
           // check axes state
           FOR #tempAxisCtr := 1 TO #MAX_NO_OF_AXES DO
             // check for axes to be existing
             IF #statAxes[#tempAxisCtr].typeOfAxis <> #AXIS_NOT_USED THEN
               // check type of axes used
               IF #statAxes[#tempAxisCtr].typeOfAxis = #TYPE_POSITIONING_AXIS THEN
                 // read TO_PositioningAxis status word
                 "LKinCtrl_GetPosAxisData"(posAxis := #statAxes[#tempAxisCtr].axis,
                                           statusWord => #statAxisStatusWord,
                                           errorDetailNumber => #statAxisErrorDetailNumber);
               ELSIF #statAxes[#tempAxisCtr].typeOfAxis = #TYPE_SYNCHRONOUS_AXIS THEN
                 // read TO_SynchronousAxis status word
                 "LKinCtrl_GetSyncAxisData"(syncAxis := #statAxes[#tempAxisCtr].axis,
                                            statusWord => #statAxisStatusWord,
                                            errorDetailNumber => #statAxisErrorDetailNumber);
               END_IF;
             END_IF;

             IF #statAxisStatusWord.%X1 = FALSE THEN
               // do nothing here, continue checks
               ;
             ELSE
               // set status
               #statStatus := #ERR_AXIS_ERROR;
               // set error bit
               #statErrorAutoCleared := TRUE;
               // write axis number to diagnostics
               #statAxisNumberDiag := #tempAxisCtr;
               // set subFunctionStatus
               #statErrorDetailNumber := #statAxisErrorDetailNumber;
               // go to error state
               #statStateMachine := #ERROR_STATE;
               EXIT;
             END_IF;

           END_FOR;

         END_REGION ENABLED_AXES


       #DISABLING_AXES: // Disabling active
         REGION DISABLING_AXES
           // set status message
           #statStatus := #STATUS_DISABLING_AXES_IN_PROGRESS;

           FOR #tempAxisCtr := 1 TO #MAX_NO_OF_AXES DO
             // check for axes to be existing
             IF #statAxes[#tempAxisCtr].typeOfAxis <> #AXIS_NOT_USED THEN
               // set execute trigger for MC_POWER
               #statEnableAxis[#tempAxisCtr] := FALSE;
             END_IF;
           END_FOR;

           // reset enabled axes counter
           #statDisabledAxesCtr := 0;
           // check for disabling to have completed successfully
           FOR #tempAxisCtr := 1 TO #MAX_NO_OF_AXES DO
             // only run code for existing axes
             IF #statAxes[#tempAxisCtr].typeOfAxis <> #AXIS_NOT_USED THEN
               // check for disabling to be done
               IF #instMC_Power[#tempAxisCtr].Status = FALSE THEN
                 // count done signals
                 #statDisabledAxesCtr += 1;
               ELSIF #instMC_Power[#tempAxisCtr].Error THEN
                 // set status
                 #statStatus := #ERR_MC_POWER;
                 // set error bit
                 #statErrorAutoCleared := TRUE;
                 // write MC_HOME errorID to diagnostics
                 #statSubfunctionStatus := #instMC_Power[#tempAxisCtr].ErrorId;
                 // write axis number to diagnostics
                 #statAxisNumberDiag := #tempAxisCtr;
                 // exit FOR loop once error is found
                 EXIT;
                 // go to error state
                 #statStateMachine := #ERROR_STATE;
               END_IF;
             END_IF;
           END_FOR;

           // check for all axes to be enabled successfully
           IF #statDisabledAxesCtr = #statExsitingAxesCtr THEN
             // set status message
             #statStatus := #STATUS_ALL_AXES_DISABLED;
             // reset variable for axesEnabled output
             #statAxesEnabled := FALSE;
             // go to next state
             #statStateMachine := #DISABLED_AXES;
           END_IF;
         END_REGION DISABLING_AXES

       #DISABLED_AXES:
         REGION DISABLED_AXES
           // when disabling is complete the bit #statDisablingCompleted must be set
           #statDisablingCompleted := TRUE;
         END_REGION DISABLED_AXES


       #ERROR_STATE:
         REGION ERROR_STATE
           // Reset axesEnabled output in case of error
           #statAxesEnabled := FALSE;
         END_REGION ERROR_STATE

       ELSE // Undefined state in state machine reached
         #statStatus := #ERR_UNDEFINED_STATE;
         #statErrorUserCleared := TRUE;
     END_CASE;
   END_REGION STATE_MACHINE


   REGION CALL_MC_POWER

     FOR #tempAxisCtr := 1 TO #MAX_NO_OF_AXES DO
       // check for axes to be existing
       IF #statAxes[#tempAxisCtr].typeOfAxis <> #AXIS_NOT_USED THEN
         // check for used axis type to call corresponding FCs
         IF #statAxes[#tempAxisCtr].typeOfAxis = #TYPE_POSITIONING_AXIS THEN
           // call MC_HOME for available positioning axes
           "LKinCtrl_CallMC_Power_PosAxis"(posAxisIn := #statAxes[#tempAxisCtr].axis,
                                           enable := #statEnableAxis[#tempAxisCtr],
                                           startMode := #startMode[#tempAxisCtr],
                                           stopMode := #stopMode[#tempAxisCtr],
                                           instMC_Power := #instMC_Power[#tempAxisCtr]);
           // check for error to be pending
           IF #instMC_Power[#tempAxisCtr].Error
             // check for no axis or kinematics errors detected prior
             AND #statStatus <> #ERR_AXIS_ERROR
             AND #statStatus <> #ERR_KIN_ERROR
           THEN
             // set status
             #statStatus := #ERR_MC_POWER;
             // set error bit
             #statErrorAutoCleared := TRUE;
             // write MC_HOME errorID to diagnostics
             #statSubfunctionStatus := #instMC_Power[#tempAxisCtr].ErrorId;
             // write axis number to diagnostics
             #statAxisNumberDiag := #tempAxisCtr;
             // exit FOR loop once error is found
             EXIT;
             // go to error state
             #statStateMachine := #ERROR_STATE;
           END_IF;

         ELSIF #statAxes[#tempAxisCtr].typeOfAxis = #TYPE_SYNCHRONOUS_AXIS THEN
           // call MC_HOME for available synchronous axes
           "LKinCtrl_CallMC_Power_SyncAxis"(syncAxisIn := #statAxes[#tempAxisCtr].axis,
                                            enable := #statEnableAxis[#tempAxisCtr],
                                            startMode := #startMode[#tempAxisCtr],
                                            stopMode := #stopMode[#tempAxisCtr],
                                            instMC_Power := #instMC_Power[#tempAxisCtr]);
           // check for error to be pending
           IF #instMC_Power[#tempAxisCtr].Error
             // check for no axis or kinematics errors detected prior
             AND #statStatus <> #ERR_AXIS_ERROR
             AND #statStatus <> #ERR_KIN_ERROR
           THEN
             // set status
             #statStatus := #ERR_MC_POWER;
             // set error bit
             #statErrorAutoCleared := TRUE;
             // write MC_HOME errorID to diagnostics
             #statSubfunctionStatus := #instMC_Power[#tempAxisCtr].ErrorId;
             // write axis number to diagnostics
             #statAxisNumberDiag := #tempAxisCtr;
             // exit FOR loop once error is found
             EXIT;
             // go to error state
             #statStateMachine := #ERROR_STATE;
           END_IF;
         END_IF;

       END_IF;
     END_FOR;

   END_REGION CALL_MC_POWER


   REGION OUTPUTS
     // Write outputs
     IF (#statDisablingCompleted = TRUE) THEN
       // Reset outputs if disabling completed
       #statBusy := FALSE;
       #statError := FALSE;
       #statErrorUserCleared := FALSE;
       #statErrorAutoCleared := FALSE;
       #statStatus := #STATUS_NO_CALL;
       #statStateMachine := #NO_PROCESSING; // Switch state machine to "no processing"

     ELSIF (#statErrorUserCleared = TRUE) AND (#statError = FALSE) THEN
       // Error can only be cleared by user; rising edge at enable input is needed to continue 
       #statBusy := FALSE;
       #statError := TRUE;
       #statStateMachine := #NO_PROCESSING; // Switch state machine to "no processing"

     ELSIF (#statErrorAutoCleared = TRUE) AND (#statError = FALSE) THEN
       // Error can be reset by FB automatically  
       #statBusy := TRUE;
       #statError := TRUE;
       // TODO: Handling of autocleared error

     ELSIF (#statErrorAutoCleared = FALSE) AND (#statErrorUserCleared = FALSE) AND (#statError = TRUE) THEN
       // If autocleared error is acknowledged
       #statBusy := TRUE;
       #statError := FALSE;
       #statStatus := #STATUS_SUBSEQUENT_CALL;
     END_IF;

     // Write static values to outputs
     #busy := #statBusy;
     #error := #statError;
     #axesEnabled := #statAxesEnabled;
     #diagnostics.status := #statStatus;
     #diagnostics.subfunctionStatus := #statSubfunctionStatus;
     #diagnostics.axisNumber := #statAxisNumberDiag;
     #diagnostics.errorDetail := #statErrorDetailNumber;
     #diagnostics.stateNumber := #statStateMachine;
   END_REGION OUTPUTS

   // =================================================================================================================
   // End of Function Block: LKinCtrl_MC_GroupPower
   // =================================================================================================================
END_FUNCTION_BLOCK

FUNCTION_BLOCK "LKinCtrl_MC_GroupHome"   // FB35022, SCL
TITLE = LKinCtrl_MC_GroupHome
{ S7_Optimized_Access := 'TRUE' }
AUTHOR : tech.team.motioncontrol@siemens.com
FAMILY : LKinCtrl
VERSION : 2.0
// FB provides funcitonalities to home all axes (TO_PositioningAxis or TO_SynchronousAxis) interconnected with TO Kinematics
   VAR_INPUT
      execute : Bool;   // Rising edge starts action once
      position : Array[1..4] of LReal;   // reference positions / orientations
      mode : Array[1..4] of Int;   // homing modes for each axis
   END_VAR
   VAR_OUTPUT
      done : Bool;   // axesGroup successfully referenced
      busy : Bool;   // FB is not finished and new output values can be expected
      active : Bool;   // FB in control of axesGroup / kinematic in motion
      commandAborted : Bool;   // command is aborted by another command
      error : Bool;   // an error occurred during the execution of the FB
      diagnostics : "LKinCtrl_typeAuxFCDiagnostics";   // diagnostics information of FB (optional)
   END_VAR
   VAR_IN_OUT
      axesGroup : TO_Kinematics;   // reference to the axesGroup
   END_VAR
   VAR
      statExecuteOld : Bool;   // Old value of 'execute' input for edge detection
      statDone : Bool;   // Static value for output 'done'
      statBusy : Bool;   // Static value for output 'busy'
      statError : Bool;   // Static value for output 'error'
      statCommandAborted : Bool;   // Static value for output 'commandAborted'
      statStatus : Word := 16#7000;   // Static value for output 'status'
      statSubfunctionStatus : Word;   // Static value for output 'subFunctionStatus'
      statAxisNumberDiag : Int;   // Static value for output 'axisNumber'
      statErrorDetailNumber : UDInt;   // static to store axis error detail number
      statStateMachine : DInt := 0;   // State in the state machine of the FB
      instMC_HOME : Array[1..4] of MC_HOME;   // multi instance array of MC_HOME
      statExecuteHoming : Array[1..4] of Bool;   // array of execute triggers for MC_HOME
      statAxes : Array[1..4] of Struct   // array of struct containing axis DB_ANY and type of axis
         typeOfAxis : Int;
         axis : DB_ANY;
      END_STRUCT;
      statHomePos : Array[1..4] of LReal;   // reference positions / orientations
      statAxisStatusWord : DWord;   // static to store axis status word
      statExsitingAxesCtr : Int;   // static counter for existing axes
      statHomedAxesCtr : Int;   // static counter for successfully homed axes
   END_VAR
   VAR_TEMP
      tempExecute : Bool;   // temporary value for input 'execute'
      tempAxisCtr : Int;   // temporary counter variable for axes
   END_VAR
   VAR CONSTANT
      FB_STATE_NO_PROCESSING : DInt := 0;   // state machine constant
      DETECT_AXES : DInt := 10;   // state machine constant
      CALC_HOME_POS : DInt := 20;   // state machine constant
      CHECK_AXES : DInt := 40;   // state machine constant
      TRIGGER_HOMING : DInt := 50;   // state machine constant
      HOMING_IN_PROGRESS : DInt := 60;   // state machine constant
      ERROR_STATE : DInt := 90;   // state machine constant
      HOMING_DONE : DInt := 100;   // state machine constant
      AXIS_NOT_USED : Int := -1;   // type of axis constant
      TYPE_POSITIONING_AXIS : Int := 0;   // type of axis constant
      TYPE_SYNCHRONOUS_AXIS : Int := 1;   // type of axis constant
      MAX_NO_OF_AXES : Int := 4;   // maximum number of axes
      STATUS_EXECUTION_FINISHED : Word := 16#0000;   // Execution finished without errors
      STATUS_NO_CALL : Word := 16#7000;   // No job being currently processed
      STATUS_FIRST_CALL : Word := 16#7001;   // First call after incoming new job (rising edge 'execute')
      STATUS_SUBSEQUENT_CALL : Word := 16#7002;   // Subsequent call during active processing without further details
      STATUS_COMMAND_ABORTED : Word := 16#7FFF;   // commanded functionality has been aborted by another command
      ERR_AXIS_ERROR : Word := 16#8350;   // error pending at axis
      ERR_MC_HOME : Word := 16#8351;   // error during execution of MC_HOME for axis
      ERR_UNDEFINED_STATE : Word := 16#8600;   // error due to an undefined state in state machine
   END_VAR
   // statAxes[1].typeOfAxis := -1;
BEGIN
   //==========================================================================================
   // SIEMENS AG
   // (c)Copyright 2019 All Rights Reserved
   //------------------------------------------------------------------------------------------
   // Library: LKinCtrl
   // Tested with: S7-1517T-3 PN/DP
   // Engineering: TIA Portal V15
   // Restrictions: ---
   // Requirements: S7-1500T FW 2.5
   // Functionality: LKinCtrl_MC_GroupHome
   // The FB is executing MC_HOME function blocks to reference all axes
   // corresponding to a specific axesGroup (TO Kinematics)
   // 
   // Support: tech.team.motioncontrol@siemens.com
   // Note: Parameter comments are only available in language 'English (United States)'
   //------------------------------------------------------------------------------------------
   // Change log table:
   // Version    Date          Expert in charge    Changes applied
   // 01.00.00   26.02.2019    JR                  First release version v1.0
   //===========================================================================================


   #tempExecute := #execute; // Work with temporary value / create process image

   REGION TRIGGERING
     IF (#tempExecute = TRUE) AND (#statExecuteOld = FALSE) // Check if FB is triggered
     THEN // First call; initialize FB
       #statDone := FALSE;
       #statBusy := TRUE;
       #statError := FALSE;
       #statStatus := #STATUS_FIRST_CALL;

       #statStateMachine := #DETECT_AXES; // State machine - start processing

       // Initialize functionality: reset of variables, diagnostics, etc.
       #statAxisStatusWord := 16#0;
       #statExsitingAxesCtr := 0;
       #statHomedAxesCtr := 0;
       #statErrorDetailNumber := 0;
       #statAxisNumberDiag := 0;
       #statSubfunctionStatus := 16#0;

       // Initialize functionality: call subsidiary FBs with FALSE
       FOR #tempAxisCtr := 1 TO #MAX_NO_OF_AXES DO
         // call all MC_HOME FBs with false
         #instMC_HOME[#tempAxisCtr].Execute := FALSE;
         // array variable resets
         #statExecuteHoming[#tempAxisCtr] := FALSE;
         #statAxes[#tempAxisCtr].axis := 0;
         #statAxes[#tempAxisCtr].typeOfAxis := #AXIS_NOT_USED;
         #statHomePos[#tempAxisCtr] := 0;
       END_FOR;


     ELSIF (#statStatus = #STATUS_FIRST_CALL) THEN
       #statStatus := #STATUS_SUBSEQUENT_CALL;
     END_IF;

     // Edge detection 'execute' input
     #statExecuteOld := #tempExecute;
   END_REGION TRIGGERING

   IF (#statStatus = #STATUS_NO_CALL) THEN
     // Nothing to do -> End here to reduce "system load"
     RETURN;
   END_IF;

   REGION STATE_MACHINE
     CASE #statStateMachine OF // State machine of FB
       #FB_STATE_NO_PROCESSING: // No processing active (Note: this state must always be present and left empty)
         ;

       #DETECT_AXES: // Processing active
         REGION DETECT_AXES
           // check available & connected axes at TO_Kinematics
           // assign DB number of connected axis to DB_ANY type
           IF #axesGroup.KinematicsAxis.A1 <> 0 THEN
             #statAxes[1].axis := #axesGroup.KinematicsAxis.A1;
             #statExsitingAxesCtr += 1;
           END_IF;
           IF #axesGroup.KinematicsAxis.A2 <> 0 THEN
             #statAxes[2].axis := #axesGroup.KinematicsAxis.A2;
             #statExsitingAxesCtr += 1;
           END_IF;
           IF #axesGroup.KinematicsAxis.A3 <> 0 THEN
             #statAxes[3].axis := #axesGroup.KinematicsAxis.A3;
             #statExsitingAxesCtr += 1;
           END_IF;
           IF #axesGroup.KinematicsAxis.A4 <> 0 THEN
             #statAxes[4].axis := #axesGroup.KinematicsAxis.A4;
             #statExsitingAxesCtr += 1;
           END_IF;

           // detect type of axis once for later call of corresponding FCs
           FOR #tempAxisCtr := 1 TO #MAX_NO_OF_AXES DO
             // check for axes to be existing
             IF #statAxes[#tempAxisCtr].axis <> 0 THEN
               IF TypeOfDB(#statAxes[#tempAxisCtr].axis) = TO_PositioningAxis THEN
                 // set type of axis to PosAxis
                 #statAxes[#tempAxisCtr].typeOfAxis := #TYPE_POSITIONING_AXIS;
               ELSIF TypeOfDB(#statAxes[#tempAxisCtr].axis) = TO_SynchronousAxis THEN
                 // set type of axis to PosAxis
                 #statAxes[#tempAxisCtr].typeOfAxis := #TYPE_SYNCHRONOUS_AXIS;
               END_IF;
             ELSE
               // set type of axis to 'not used'
               #statAxes[#tempAxisCtr].typeOfAxis := #AXIS_NOT_USED;
             END_IF;

           END_FOR;


           // go to next state
           #statStateMachine := #CALC_HOME_POS;
         END_REGION DETECT_AXES


       #CALC_HOME_POS:
         REGION CALC_HOME_POS
           // calculations for homing positions according to coordSystem added later
           #statHomePos := #position;

           // go to next state
           #statStateMachine := #CHECK_AXES;
         END_REGION CALC_HOME_POS


       #CHECK_AXES:
         REGION CHECK_AXES
           FOR #tempAxisCtr := 1 TO #MAX_NO_OF_AXES DO
             // check for axes to be existing
             IF #statAxes[#tempAxisCtr].typeOfAxis <> #AXIS_NOT_USED THEN
               // check type of axes used
               IF #statAxes[#tempAxisCtr].typeOfAxis = #TYPE_POSITIONING_AXIS THEN
                 // read TO_PositioningAxis status word
                 "LKinCtrl_GetPosAxisData"(posAxis := #statAxes[#tempAxisCtr].axis,
                                           statusWord => #statAxisStatusWord,
                                           errorDetailNumber=> #statErrorDetailNumber);
               ELSIF #statAxes[#tempAxisCtr].typeOfAxis = #TYPE_SYNCHRONOUS_AXIS THEN
                 // read TO_SynchronousAxis status word
                 "LKinCtrl_GetSyncAxisData"(syncAxis := #statAxes[#tempAxisCtr].axis,
                                            statusWord => #statAxisStatusWord,
                                            errorDetailNumber=> #statErrorDetailNumber);
               END_IF;
             END_IF;

             IF #statAxisStatusWord.%X1 = FALSE THEN
               // do nothing here, continue axes checks
               ;
             ELSE
               #statStatus := #ERR_AXIS_ERROR;
               // write axis number to diagnostics
               #statAxisNumberDiag := #tempAxisCtr;
               // go to error state
               #statStateMachine := #ERROR_STATE;
               EXIT;
             END_IF;

           END_FOR;

           // check for no error to be pending
           IF #statStatus.%X15 = FALSE THEN
             // go to next state
             #statStateMachine := #TRIGGER_HOMING;
           END_IF;
         END_REGION CHECK_AXES



       #TRIGGER_HOMING: // execute homing procedure
         REGION TRIGGER_HOMING
           FOR #tempAxisCtr := 1 TO #MAX_NO_OF_AXES DO
             // check for axes to be existing
             IF #statAxes[#tempAxisCtr].typeOfAxis <> #AXIS_NOT_USED THEN
               // set execute trigger for MC_HOME
               #statExecuteHoming[#tempAxisCtr] := TRUE;
             END_IF;
           END_FOR;

           // go to next state
           #statStateMachine := #HOMING_IN_PROGRESS;
         END_REGION TRIGGER_HOMING


       #HOMING_IN_PROGRESS:
         REGION HOMING_IN_PROGRESS
           // reset homed axes counter
           #statHomedAxesCtr := 0;
           // check for homing to have completed successfully
           FOR #tempAxisCtr := 1 TO #MAX_NO_OF_AXES DO
             // only run code for existing axes
             IF #statAxes[#tempAxisCtr].typeOfAxis <> #AXIS_NOT_USED THEN
               // check for homing to be done
               IF #instMC_HOME[#tempAxisCtr].Done THEN
                 // count done signals
                 #statHomedAxesCtr += 1;

               ELSIF #instMC_HOME[#tempAxisCtr].CommandAborted THEN
                 // set status
                 #statStatus := #STATUS_COMMAND_ABORTED;
                 // write MC_HOME errorID to diagnostics
                 #statSubfunctionStatus := #instMC_HOME[#tempAxisCtr].ErrorId;
                 // write axis number to diagnostics
                 #statAxisNumberDiag := #tempAxisCtr;
                 // exit FOR loop once error is found
                 EXIT;

               ELSIF #instMC_HOME[#tempAxisCtr].Error THEN
                 // set status
                 #statStatus := #ERR_MC_HOME;
                 // write MC_HOME errorID to diagnostics
                 #statSubfunctionStatus := #instMC_HOME[#tempAxisCtr].ErrorId;
                 // write axis number to diagnostics
                 #statAxisNumberDiag := #tempAxisCtr;
                 // exit FOR loop once error is found
                 EXIT;
                 // go to error state
                 #statStateMachine := #ERROR_STATE;
               END_IF;
             END_IF;
           END_FOR;

           // check for all axes to be homed successfully
           IF #statHomedAxesCtr = #statExsitingAxesCtr THEN
             FOR #tempAxisCtr := 1 TO #MAX_NO_OF_AXES DO
               // reset execute trigger for MC_HOME
               #statExecuteHoming[#tempAxisCtr] := FALSE;
             END_FOR;

             // go to next state
             #statStateMachine := #HOMING_DONE;
           END_IF;
         END_REGION HOMING_IN_PROGRESS


       #HOMING_DONE:
         REGION HOMING_DONE
           // set status to initiate end of FB execution
           #statStatus := #STATUS_EXECUTION_FINISHED;

         END_REGION HOMING_DONE


       #ERROR_STATE:
         // do nothing
         ;

       ELSE // Undefined state in state machine reached
         #statStatus := #ERR_UNDEFINED_STATE;
     END_CASE;
   END_REGION STATE_MACHINE

   REGION CALL_MC_HOME
     FOR #tempAxisCtr := 1 TO #MAX_NO_OF_AXES DO
       // check for axes to be existing
       IF #statAxes[#tempAxisCtr].typeOfAxis <> #AXIS_NOT_USED THEN
         // check for used axis type to call corresponding FCs
         IF #statAxes[#tempAxisCtr].typeOfAxis = #TYPE_POSITIONING_AXIS THEN
           // call MC_HOME for available positioning axes
           "LKinCtrl_CallMC_Home_PosAxis"(posAxisIn := #statAxes[#tempAxisCtr].axis,
                                          execute := #statExecuteHoming[#tempAxisCtr],
                                          position := #statHomePos[#tempAxisCtr],
                                          mode := #mode[#tempAxisCtr],
                                          instMC_Home := #instMC_HOME[#tempAxisCtr]);
         ELSIF #statAxes[#tempAxisCtr].typeOfAxis = #TYPE_SYNCHRONOUS_AXIS THEN
           // call MC_HOME for available synchronous axes
           "LKinCtrl_CallMC_Home_SyncAxis"(syncAxisIn := #statAxes[#tempAxisCtr].axis,
                                           execute := #statExecuteHoming[#tempAxisCtr],
                                           position := #statHomePos[#tempAxisCtr],
                                           mode := #mode[#tempAxisCtr],
                                           instMC_Home := #instMC_HOME[#tempAxisCtr]);
         END_IF;

       END_IF;
     END_FOR;


   END_REGION


   REGION OUTPUTS
     // Write outputs
     IF (#statStatus = #STATUS_EXECUTION_FINISHED) AND (#statDone = FALSE) THEN // Execution finished without errors
       #statDone := TRUE;
       #statBusy := FALSE;
       #statError := FALSE;
       #statStateMachine := #FB_STATE_NO_PROCESSING; // Switch state machine to "no processing"

     ELSIF (#statStatus.%X15 = TRUE) AND (#statError = FALSE) THEN // Error occurred (#statStatus is 16#8000 to 16#FFFF)
       #statDone := FALSE;
       #statBusy := FALSE;
       #statError := TRUE;
       #statStateMachine := #FB_STATE_NO_PROCESSING; // Switch state machine to "no processing"

     ELSIF (#tempExecute = FALSE) AND ((#statDone = TRUE) OR (#statError = TRUE)) THEN // Reset outputs
       #statDone := FALSE;
       #statBusy := FALSE;
       #statError := FALSE;
       #statStatus := #STATUS_NO_CALL;
       // TODO: Reset application specific outputs
     END_IF;

     // Write static values to outputs
     #done := #statDone;
     #busy := #statBusy;
     #error := #statError;
     #diagnostics.status := #statStatus;
     #diagnostics.subfunctionStatus := #statSubfunctionStatus;
     #diagnostics.axisNumber := #statAxisNumberDiag;
     #diagnostics.errorDetail := #statErrorDetailNumber;
     #diagnostics.stateNumber := #statStateMachine;
     // TODO: Write application specific static values to outputs
   END_REGION OUTPUTS

   // =================================================================================================================
   // End of Function Block: LKinCtrl_MC_GroupHome
   // =================================================================================================================
END_FUNCTION_BLOCK

FUNCTION_BLOCK "LKinCtrl_MC_GroupReset"   // FB35023, SCL
TITLE = LKinCtrl_MC_GroupReset
{ S7_Optimized_Access := 'TRUE' }
AUTHOR : tech.team.motioncontrol@siemens.com
FAMILY : LKinCtrl
VERSION : 2.0
// FB provides funcitonalities to reset all axes (TO_PositioningAxis or TO_SynchronousAxis) interconnected with TO Kinematics and the TO Kinematics itself using internal MC_RESET
   VAR_INPUT
      execute : Bool;   // Rising edge starts action once
      restart : Array[1..5] of Bool;   // reinitialization of technology object
   END_VAR
   VAR_OUTPUT
      done : Bool;   // axesGroup successfully referenced
      busy : Bool;   // FB is not finished and new output values can be expected
      active : Bool;   // FB in control of axesGroup / kinematic in motion
      commandAborted : Bool;   // command is aborted by another command
      error : Bool;   // an error occurred during the execution of the FB
      diagnostics : "LKinCtrl_typeAuxFCDiagnostics";   // diagnostics information of FB (optional)
   END_VAR
   VAR_IN_OUT
      axesGroup : TO_Kinematics;   // reference to the axesGroup
   END_VAR
   VAR
      statExecuteOld : Bool;   // Old value of 'execute' input for edge detection
      statDone : Bool;   // Static value for output 'done'
      statBusy : Bool;   // Static value for output 'busy'
      statError : Bool;   // Static value for output 'error'
      statStatus : Word := 16#7000;   // Static value for output 'status'
      statSubfunctionStatus : Word;   // Static value for output 'subFunctionStatus'
      statAxisNumberDiag : Int;   // Static value for output 'axisNumber'
      statErrorDetailNumber : UDInt;   // static to store axis error detail number
      statStateMachine : DInt := 0;   // State in the state machine of the FB
      instMC_RESET_Axes : Array[1..#MAX_NO_OF_AXES] of MC_RESET;   // multi instance array of MC_RESET for axes
      instMC_RESET_Kin : MC_RESET;   // multi instance of MC_RESET for TO_Kinematics
      statExecuteResetAxis : Array[1..#MAX_NO_OF_AXES] of Bool;   // array of execute triggers for MC_HOME
      statExecuteResetKin : Bool;   // execute trigger for TO_Kinematics
      statAxes : Array[1..#MAX_NO_OF_AXES] of Struct   // array of struct containing axis DB_ANY and type of axis
         typeOfAxis : Int;
         axis : DB_ANY;
      END_STRUCT;
      statAxisStatusWord : DWord;   // static to store axis status word
      statExsitingAxesCtr : Int;   // static counter for existing axes
      statResetAxesCtr : Int;   // static counter for successfully homed axes
   END_VAR
   VAR_TEMP
      tempExecute : Bool;   // temporary value for input 'execute'
      tempAxisCtr : Int;   // temporary counter variable for axes
   END_VAR
   VAR CONSTANT
      NO_PROCESSING : DInt := 0;   // state machine constant
      DETECT_AXES : DInt := 10;   // state machine constant
      CALC_HOME_POS : DInt := 20;   // state machine constant
      CHECK_AXES : DInt := 40;   // state machine constant
      TRIGGER_RESET : DInt := 50;   // state machine constant
      RESETTING_IN_PROGRESS : DInt := 60;   // state machine constant
      ERROR_STATE : DInt := 90;   // state machine constant
      RESETTING_DONE : DInt := 100;   // state machine constant
      AXIS_NOT_USED : Int := -1;   // type of axis constant
      TYPE_POSITIONING_AXIS : Int := 0;   // type of axis constant
      TYPE_SYNCHRONOUS_AXIS : Int := 1;   // type of axis constant
      TYPE_TO_KINEMATICS : Int := 2;   // type of axis constant
      MAX_NO_OF_AXES : Int := 4;   // maximum number of axes
      STATUS_EXECUTION_FINISHED : Word := 16#0000;   // Execution finished without errors
      STATUS_NO_CALL : Word := 16#7000;   // No job being currently processed
      STATUS_FIRST_CALL : Word := 16#7001;   // First call after incoming new job (rising edge 'execute')
      STATUS_SUBSEQUENT_CALL : Word := 16#7002;   // Subsequent call during active processing without further details
      STATUS_COMMAND_ABORTED : Word := 16#7FFF;   // Commanded functionality has been aborted by another command
      ERR_AXIS_ERROR : Word := 16#8360;   // error pending at axis
      ERR_KIN_ERROR : Word := 16#8361;   // error pending at kinematics
      ERR_MC_RESET_AXES : Word := 16#8362;   // error during execution of MC_RESET for axis
      ERR_MC_RESET_KIN : Word := 16#8363;   // error during execution of MC_RESET for kinematics
      ERR_UNDEFINED_STATE : Word := 16#8600;   // error due to an undefined state in state machine
   END_VAR
   // statAxes[1].typeOfAxis := -1;
BEGIN
   //==========================================================================================
   // SIEMENS AG
   // (c)Copyright 2019 All Rights Reserved
   //------------------------------------------------------------------------------------------
   // Library: LKinCtrl
   // Tested with: S7-1517T-3 PN/DP
   // Engineering: TIA Portal V15
   // Restrictions: ---
   // Requirements: S7-1500T FW 2.5
   // Functionality: LKinCtrl_MC_GroupReset
   // The FB is executing MC_RESET function blocks to reset all axes
   // and the axesGroup (TO Kinematics)
   // 
   // Support: tech.team.motioncontrol@siemens.com
   // Note: Parameter comments are only available in language 'English (United States)'
   //------------------------------------------------------------------------------------------
   // Change log table:
   // Version    Date          Expert in charge    Changes applied
   // 01.00.00   27.02.2019    JR                  First release version v1.0
   //===========================================================================================

   #tempExecute := #execute; // Work with temporary value / create process image

   REGION TRIGGERING
     IF (#tempExecute = TRUE) AND (#statExecuteOld = FALSE) // Check if FB is triggered
     THEN // First call; initialize FB
       #statDone := FALSE;
       #statBusy := TRUE;
       #statError := FALSE;
       #statStatus := #STATUS_FIRST_CALL;

       #statStateMachine := #DETECT_AXES; // State machine - start processing

       // Initialize functionality: reset of variables, diagnostics, etc.
       #statAxisStatusWord := 16#0;
       #statExsitingAxesCtr := 0;
       #statResetAxesCtr := 0;
       #statErrorDetailNumber := 0;
       #statAxisNumberDiag := 0;
       #statSubfunctionStatus := 16#0;

       // Initialize functionality: call subsidiary FBs with FALSE
       FOR #tempAxisCtr := 1 TO #MAX_NO_OF_AXES DO
         // call all MC_HOME FBs with false
         #instMC_RESET_Axes[#tempAxisCtr].Execute := FALSE;
         // array variable resets
         #statExecuteResetAxis[#tempAxisCtr] := FALSE;
         #statAxes[#tempAxisCtr].axis := 0;
         #statAxes[#tempAxisCtr].typeOfAxis := #AXIS_NOT_USED;
       END_FOR;


     ELSIF (#statStatus = #STATUS_FIRST_CALL) THEN
       #statStatus := #STATUS_SUBSEQUENT_CALL;
     END_IF;

     // Edge detection 'execute' input
     #statExecuteOld := #tempExecute;
   END_REGION TRIGGERING

   IF (#statStatus = #STATUS_NO_CALL) THEN
     // Nothing to do -> End here to reduce "system load"
     RETURN;
   END_IF;

   REGION STATE_MACHINE
     CASE #statStateMachine OF // State machine of FB
       #NO_PROCESSING: // No processing active (Note: this state must always be present and left empty)
         ;

       #DETECT_AXES: // Processing active
         REGION DETECT_AXES
           // check available & connected axes at TO_Kinematics
           // assign DB number of connected axis to DB_ANY type
           IF #axesGroup.KinematicsAxis.A1 <> 0 THEN
             #statAxes[1].axis := #axesGroup.KinematicsAxis.A1;
             #statExsitingAxesCtr += 1;
           END_IF;
           IF #axesGroup.KinematicsAxis.A2 <> 0 THEN
             #statAxes[2].axis := #axesGroup.KinematicsAxis.A2;
             #statExsitingAxesCtr += 1;
           END_IF;
           IF #axesGroup.KinematicsAxis.A3 <> 0 THEN
             #statAxes[3].axis := #axesGroup.KinematicsAxis.A3;
             #statExsitingAxesCtr += 1;
           END_IF;
           IF #axesGroup.KinematicsAxis.A4 <> 0 THEN
             #statAxes[4].axis := #axesGroup.KinematicsAxis.A4;
             #statExsitingAxesCtr += 1;
           END_IF;

           // detect type of axis once for later call of corresponding FCs
           FOR #tempAxisCtr := 1 TO #MAX_NO_OF_AXES DO
             // check for axes to be existing
             IF #statAxes[#tempAxisCtr].axis <> 0 THEN
               IF TypeOfDB(#statAxes[#tempAxisCtr].axis) = TO_PositioningAxis THEN
                 // set type of axis to PosAxis
                 #statAxes[#tempAxisCtr].typeOfAxis := #TYPE_POSITIONING_AXIS;
               ELSIF TypeOfDB(#statAxes[#tempAxisCtr].axis) = TO_SynchronousAxis THEN
                 // set type of axis to PosAxis
                 #statAxes[#tempAxisCtr].typeOfAxis := #TYPE_SYNCHRONOUS_AXIS;
               END_IF;
             ELSE
               // set type of axis to 'not used'
               #statAxes[#tempAxisCtr].typeOfAxis := #AXIS_NOT_USED;
             END_IF;

           END_FOR;


           // go to next state
           #statStateMachine := #TRIGGER_RESET;
         END_REGION DETECT_AXES

       #TRIGGER_RESET: // execute homing procedure
         REGION TRIGGER_RESET
           FOR #tempAxisCtr := 1 TO #MAX_NO_OF_AXES DO
             // check for axes to be existing
             IF #statAxes[#tempAxisCtr].typeOfAxis <> #AXIS_NOT_USED THEN
               // set execute trigger for MC_RESET
               #statExecuteResetAxis[#tempAxisCtr] := TRUE;
             END_IF;
           END_FOR;
           // set execute trigger for TO_Kinematics
           #statExecuteResetKin := TRUE;

           // go to next state
           #statStateMachine := #RESETTING_IN_PROGRESS;
         END_REGION TRIGGER_RESET

       #RESETTING_IN_PROGRESS:
         REGION RESETTING_IN_PROGRESS
           // reset homed axes counter
           #statResetAxesCtr := 0;
           // check for homing to have completed successfully
           FOR #tempAxisCtr := 1 TO #MAX_NO_OF_AXES DO
             // only run code for existing axes
             IF #statAxes[#tempAxisCtr].typeOfAxis <> #AXIS_NOT_USED THEN
               // check for homing to be done
               IF #instMC_RESET_Axes[#tempAxisCtr].Done THEN
                 // count done signals
                 #statResetAxesCtr += 1;

               ELSIF #instMC_RESET_Axes[#tempAxisCtr].CommandAborted THEN
                 // set status
                 #statStatus := #STATUS_COMMAND_ABORTED;
                 // write MC_RESET errorID to diagnostics
                 #statSubfunctionStatus := #instMC_RESET_Axes[#tempAxisCtr].ErrorId;
                 // write axis number to diagnostics
                 #statAxisNumberDiag := #tempAxisCtr;
                 // exit FOR loop once error is found
                 EXIT;

               ELSIF #instMC_RESET_Axes[#tempAxisCtr].Error THEN
                 // set status
                 #statStatus := #ERR_MC_RESET_AXES;
                 // write MC_HOME errorID to diagnostics
                 #statSubfunctionStatus := #instMC_RESET_Axes[#tempAxisCtr].ErrorId;
                 // write axis number to diagnostics
                 #statAxisNumberDiag := #tempAxisCtr;
                 // exit FOR loop once error is found
                 EXIT;
                 // go to error state
                 #statStateMachine := #ERROR_STATE;
               END_IF;
             END_IF;
           END_FOR;

           // check for TO Kinematics reset to be completed
           IF #instMC_RESET_Kin.Done THEN
             // count done signals
             #statResetAxesCtr += 1;

           ELSIF #instMC_RESET_Kin.#CommandAborted THEN
             // set status
             #statStatus := #STATUS_COMMAND_ABORTED;
             // write MC_RESET errorID to diagnostics
             #statSubfunctionStatus := #instMC_RESET_Kin.ErrorId;
             // write axis number to diagnostics
             #statAxisNumberDiag := #MAX_NO_OF_AXES + 1;

           ELSIF #instMC_RESET_Kin.#Error THEN
             // set status
             #statStatus := #ERR_MC_RESET_KIN;
             // write MC_HOME errorID to diagnostics
             #statSubfunctionStatus := #instMC_RESET_Kin.ErrorId;
             // write axis number to diagnostics
             #statAxisNumberDiag := #MAX_NO_OF_AXES + 1;
             // go to error state
             #statStateMachine := #ERROR_STATE;
           END_IF;


           // check for all axes (+ TO_Kinematics) to be homed successfully
           IF #statResetAxesCtr = #statExsitingAxesCtr + 1 THEN
             FOR #tempAxisCtr := 1 TO #MAX_NO_OF_AXES DO
               // reset execute trigger for MC_RESET for axes
               #statExecuteResetAxis[#tempAxisCtr] := FALSE;
               // reset execute trigger for MC_RESET for TO_Kinematics
               #statExecuteResetKin := FALSE;
             END_FOR;

             // go to next state
             #statStateMachine := #CHECK_AXES;
           ELSE
             ;
           END_IF;
         END_REGION RESETTING_IN_PROGRESS

       #CHECK_AXES:
         REGION CHECK_AXES
           FOR #tempAxisCtr := 1 TO #MAX_NO_OF_AXES DO
             // check for axes to be existing
             IF #statAxes[#tempAxisCtr].typeOfAxis <> #AXIS_NOT_USED THEN
               // check type of axes used
               IF #statAxes[#tempAxisCtr].typeOfAxis = #TYPE_POSITIONING_AXIS THEN
                 // read TO_PositioningAxis status word
                 "LKinCtrl_GetPosAxisData"(posAxis := #statAxes[#tempAxisCtr].axis,
                                           statusWord => #statAxisStatusWord,
                                           errorDetailNumber=> #statErrorDetailNumber);
               ELSIF #statAxes[#tempAxisCtr].typeOfAxis = #TYPE_SYNCHRONOUS_AXIS THEN
                 // read TO_SynchronousAxis status word
                 "LKinCtrl_GetSyncAxisData"(syncAxis := #statAxes[#tempAxisCtr].axis,
                                            statusWord => #statAxisStatusWord,
                                            errorDetailNumber=> #statErrorDetailNumber);
               END_IF;
             END_IF;

             IF #statAxisStatusWord.%X1 = FALSE THEN
               // do nothing here, continue checks
               ;
             ELSE
               #statStatus := #ERR_AXIS_ERROR;
               // write axis number to diagnostics
               #statAxisNumberDiag := #tempAxisCtr;
               // go to error state
               #statStateMachine := #ERROR_STATE;
               EXIT;
             END_IF;

           END_FOR;

           // check TO_Kinematics to have no errors pending
           IF #axesGroup.StatusWord.%X1 = FALSE THEN
             // do nothing here, continue checks
             ;
           ELSE
             #statStatus := #ERR_KIN_ERROR;
             // go to error state
             #statStateMachine := #ERROR_STATE;
           END_IF;


           // check for no error to be pending
           IF #statStatus.%X15 = FALSE THEN
             // go to next state
             #statStateMachine := #RESETTING_DONE;
           END_IF;
         END_REGION CHECK_AXES



       #RESETTING_DONE:
         REGION RESETTING_DONE
           // set status to initiate end of FB execution
           #statStatus := #STATUS_EXECUTION_FINISHED;

         END_REGION RESETTING_DONE


       #ERROR_STATE:
         // do nothing
         ;

       ELSE // Undefined state in state machine reached
         #statStatus := #ERR_UNDEFINED_STATE;
     END_CASE;

   END_REGION STATE_MACHINE


   REGION CALL_MC_RESET

     FOR #tempAxisCtr := 1 TO #MAX_NO_OF_AXES DO
       // check for axes to be existing
       IF #statAxes[#tempAxisCtr].typeOfAxis <> #AXIS_NOT_USED THEN
         // check for used axis type to call corresponding FCs
         IF #statAxes[#tempAxisCtr].typeOfAxis = #TYPE_POSITIONING_AXIS THEN
           // call MC_HOME for available positioning axes
           "LKinCtrl_CallMC_Reset_PosAxis"(posAxisIn := #statAxes[#tempAxisCtr].axis,
                                           execute := #statExecuteResetAxis[#tempAxisCtr],
                                           restart := #restart[#tempAxisCtr],
                                           instMC_Reset := #instMC_RESET_Axes[#tempAxisCtr]);
         ELSIF #statAxes[#tempAxisCtr].typeOfAxis = #TYPE_SYNCHRONOUS_AXIS THEN
           // call MC_HOME for available synchronous axes
           "LKinCtrl_CallMC_Reset_SyncAxis"(syncAxisIn := #statAxes[#tempAxisCtr].axis,
                                            execute := #statExecuteResetAxis[#tempAxisCtr],
                                            restart := #restart[#tempAxisCtr],
                                            instMC_Reset := #instMC_RESET_Axes[#tempAxisCtr]);
         END_IF;

       END_IF;
     END_FOR;
     #instMC_RESET_Kin(Axis := #axesGroup,
                       Execute := #statExecuteResetKin,
                       Restart := #restart[#MAX_NO_OF_AXES + 1]); 

   END_REGION CALL_MC_RESET


   REGION OUTPUTS
     // Write outputs
     IF (#statStatus = #STATUS_EXECUTION_FINISHED) AND (#statDone = FALSE) THEN // Execution finished without errors
       #statDone := TRUE;
       #statBusy := FALSE;
       #statError := FALSE;
       #statStateMachine := #NO_PROCESSING; // Switch state machine to "no processing"

     ELSIF (#statStatus.%X15 = TRUE) AND (#statError = FALSE) THEN // Error occurred (#statStatus is 16#8000 to 16#FFFF)
       #statDone := FALSE;
       #statBusy := FALSE;
       #statError := TRUE;
       #statStateMachine := #NO_PROCESSING; // Switch state machine to "no processing"

     ELSIF (#tempExecute = FALSE) AND ((#statDone = TRUE) OR (#statError = TRUE)) THEN // Reset outputs
       #statDone := FALSE;
       #statBusy := FALSE;
       #statError := FALSE;
       #statStatus := #STATUS_NO_CALL;
       // TODO: Reset application specific outputs
     END_IF;

     // Write static values to outputs
     #done := #statDone;
     #busy := #statBusy;
     #error := #statError;
     #diagnostics.status := #statStatus;
     #diagnostics.subfunctionStatus := #statSubfunctionStatus;
     #diagnostics.axisNumber := #statAxisNumberDiag;
     #diagnostics.errorDetail := #statErrorDetailNumber;
     #diagnostics.stateNumber := #statStateMachine;
   END_REGION OUTPUTS

   // =================================================================================================================
   // End of Function Block: LKinCtrl_MC_GroupReset
   // =================================================================================================================
END_FUNCTION_BLOCK

// folder: LKinCtrl_Blocks/LKinCtrl_AuxBlocks/LKinCtrl_AuxSubBlocks

FUNCTION "LKinCtrl_GetPosAxisData" : Void   // FC35021, SCL
{ S7_Optimized_Access := 'TRUE' }
VERSION : 0.1
   VAR_INPUT
      posAxis : TO_PositioningAxis;   // PositioningAxis to get data from
   END_VAR
   VAR_OUTPUT
      statusWord : DWord;   // axis status word
      errorDetailNumber : UDInt;   // axis error detail number
   END_VAR
BEGIN
   //================================================================================
   // SIEMENS AG
   // (c)Copyright 2019 All Rights Reserved
   //--------------------------------------------------------------------------------
   // Library: LKinCtrl
   // Tested with: S7-1517T-3 PN
   // Engineering: TIA Portal V15
   // Restrictions: -
   // Requirements: S7-1500T FW 2.5
   // Functionality: Get PositiongAxis StatusWord
   // Support: tech.team.motioncontrol@siemens.com
   // Note: Parameter comments are only available in language 'English (United States)'
   //-----------------------------------------------------------------------------
   // Change log table:
   // Version    Date          Expert in charge    Changes applied
   // 01.00.00   27.02.2019    JR                  First released version
   //===========================================================================================

   // return statusWord of PositioningAxis
   #statusWord := #posAxis.StatusWord;
   // check for error to be pending
   IF #statusWord.%X1 THEN
     // return error detail number
     #errorDetailNumber := #posAxis.ErrorDetail.Number;
   END_IF;
END_FUNCTION

FUNCTION "LKinCtrl_GetSyncAxisData" : Void   // FC35022, SCL
{ S7_Optimized_Access := 'TRUE' }
VERSION : 0.1
   VAR_INPUT
      syncAxis : TO_SynchronousAxis;   // SynchronousAxis to get data from
   END_VAR
   VAR_OUTPUT
      statusWord : DWord;   // axis status word
      errorDetailNumber : UDInt;   // axis error detail number
   END_VAR
BEGIN
   //================================================================================
   // SIEMENS AG
   // (c)Copyright 2019 All Rights Reserved
   //--------------------------------------------------------------------------------
   // Library: LKinCtrl
   // Tested with: S7-1517T-3 PN
   // Engineering: TIA Portal V15
   // Restrictions: -
   // Requirements: S7-1500T FW 2.5
   // Functionality: Get PositiongAxis StatusWord
   // Support: tech.team.motioncontrol@siemens.com
   // Note: Parameter comments are only available in language 'English (United States)'
   //-----------------------------------------------------------------------------
   // Change log table:
   // Version    Date          Expert in charge    Changes applied
   // 01.00.00   27.02.2019    JR                  First released version
   //===========================================================================================

   // return statusWord of SynchronousAxis
   #statusWord := #syncAxis.StatusWord;
   // check for error to be pending
   IF #statusWord.%X1 THEN
     // return error detail number
     #errorDetailNumber := #syncAxis.ErrorDetail.Number;
   END_IF;
END_FUNCTION

FUNCTION "LKinCtrl_CallMC_Home_PosAxis" : Void   // FC35023, SCL
{ S7_Optimized_Access := 'TRUE' }
VERSION : 0.1
   VAR_INPUT
      posAxisIn : TO_PositioningAxis;   // PositioningAxis to access
      execute : Bool;   // execute trigger
      position : LReal;   // home position
      mode : Int;   // homing mode
   END_VAR
   VAR_IN_OUT
      instMC_Home : MC_HOME;   // multi instance MC_HOME
   END_VAR
BEGIN
   //================================================================================
   // SIEMENS AG
   // (c)Copyright 2019 All Rights Reserved
   //--------------------------------------------------------------------------------
   // Library: LKinCtrl
   // Tested with: S7-1517T-3 PN
   // Engineering: TIA Portal V15
   // Restrictions: -
   // Requirements: S7-1500T FW 2.5
   // Functionality: Call MC_Home
   // Support: tech.team.motioncontrol@siemens.com
   // Note: Parameter comments are only available in language 'English (United States)'
   //-----------------------------------------------------------------------------
   // Change log table:
   // Version    Date          Expert in charge    Changes applied
   // 01.00.00   27.02.2019    JR                  First released version
   //===========================================================================================

   // call MC_Home
   #instMC_Home(Axis:=#posAxisIn,
                Execute:=#execute,
                Position:=#position,
                Mode:=#mode);
END_FUNCTION

